(* Logix 5000 project; controller Seperator 1756-L85E rev 33.11; software revision 33.01; part 7 of 7 *)
(* tags used below, declared in another part *)
   Aborted : SFC_STEP;
   Aborting : SFC_STEP;
   Auto_Manual : BOOL;
   CV1 : REAL;
   CV2 : REAL;
   CV3 : DINT;
   Equilibrating : SFC_STEP;
   FI101 : REAL;
   FI102 : REAL;
   FillerPUD1 : RampUpDn;
   FillerPUD2 : RampUpDn;
   FillerPUD3 : RampUpDn;
   FillerPUD4 : RampUpDn;
   FillerPUD5 : RampUpDn;
   FillerPUD6 : RampUpDn;
   FillerPUD7 : RampUpDn;
   Filling : SFC_STEP;
   Flushing : SFC_STEP;
   Half_Sec_PLs : TIMER;
   Holding : SFC_STEP;
   Idle : SFC_STEP;
   II101 : REAL;
   Led_Code : INT;
   LevelUD1 : RampUpDn;
   LI101 : REAL;
   Main_Sequencer : DINT;
   MyP_Motor : P_Motor;   // My (Single-Speed, Non-Reversing) Motor
   PI102 : REAL;
   Qtr_Sec_PLs : TIMER;
   Random : AOI_SIM_RNG_Simple;
   Restarting : SFC_STEP;
   Sec_PLs : TIMER;
   Seperating : SFC_STEP;
   Seperator_Control : PHASE;
   Speeding : SFC_STEP;
   Starting : SFC_STEP;
   Status_Code : INT;
   Stopped : SFC_STEP;
   Stopping : SFC_STEP;
   T1 : FBD_TIMER;
   TI101 : REAL;
   TI101_Temperature : REAL;
   TI101_Temperature_PID_CV : REAL;
   TI101_Temperature_PID_PV : REAL;
   TI101_Temperature_PID_SP : REAL;
   VI101 : REAL;
(* Main_Sequencer, continued *)

ROUTINE Main_Sequencer   (* ladder *)
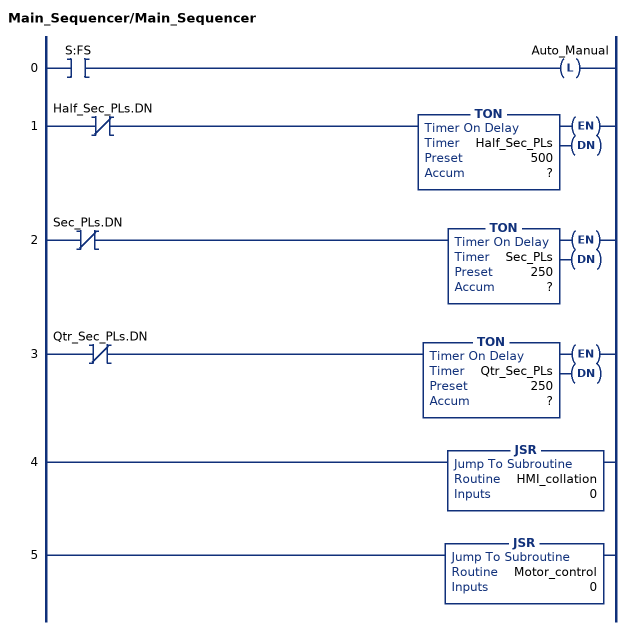
   0: XIC(S:FS)OTL(Auto_Manual);
   1: XIO(Half_Sec_PLs.DN)TON(Half_Sec_PLs,?,?);
   2: XIO(Sec_PLs.DN)TON(Sec_PLs,?,?);
   3: XIO(Qtr_Sec_PLs.DN)TON(Qtr_Sec_PLs,?,?);
   4: JSR(HMI_collation,0);
   5: JSR(Motor_control,0);
END_ROUTINE

ROUTINE Motor_control   (* ladder *)
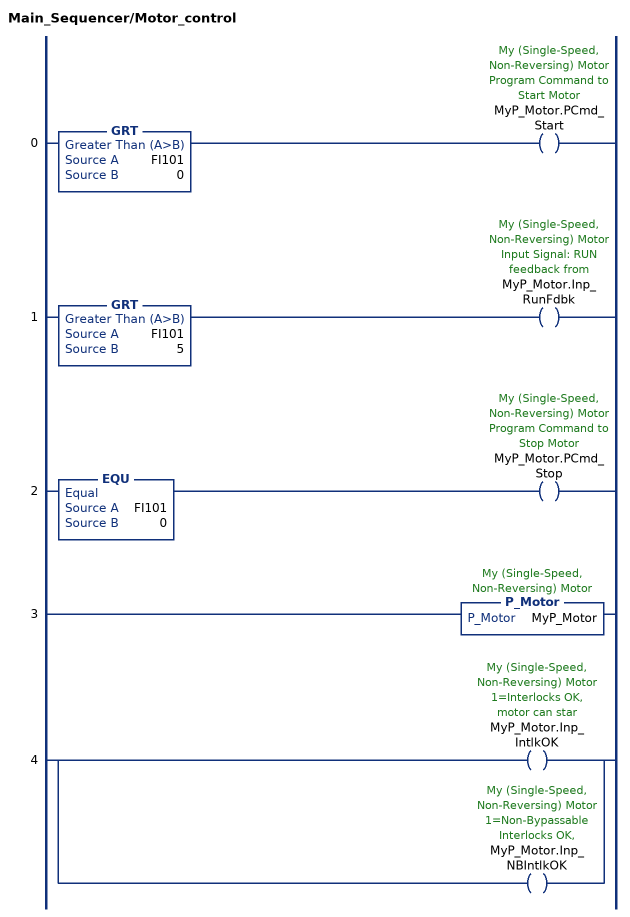
   0: GRT(FI101,0)OTE(MyP_Motor.PCmd_Start);
   1: GRT(FI101,5)OTE(MyP_Motor.Inp_RunFdbk);
   2: EQU(FI101,0)OTE(MyP_Motor.PCmd_Stop);
   3: P_Motor(MyP_Motor);
   4: [OTE(MyP_Motor.Inp_IntlkOK) ,OTE(MyP_Motor.Inp_NBIntlkOK) ];
END_ROUTINE
END_PROGRAM

PROGRAM RandomProgram   (* main routine RandomRoutine *)
VAR
   fsn : REAL := 0.19112337;
END_VAR

ROUTINE RandomRoutine   (* ladder *)
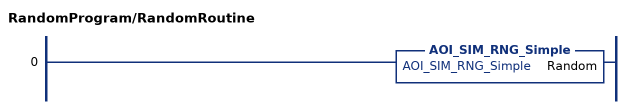
   0: AOI_SIM_RNG_Simple(Random);
END_ROUTINE
END_PROGRAM

PROGRAM RandomUpDown   (* main routine main *)
VAR
   dice001 : AOI_SIM_RNG_Simple := (Seed := 521288629, Count := 470, Number := 0.55877805);
   mult : REAL := 0.025;
   signal : REAL := 0.8641962;
   up : BOOL := 1;
END_VAR

ROUTINE main   (* ladder *)
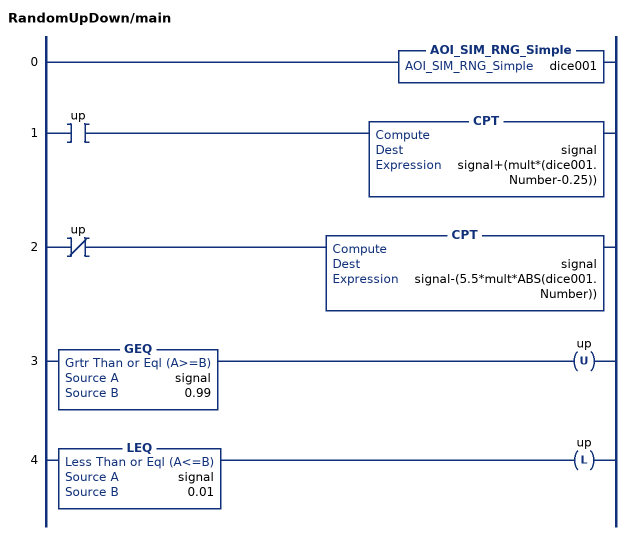
   0: AOI_SIM_RNG_Simple(dice001);
   1: XIC(up)CPT(signal,signal+(mult*(dice001.Number-0.25)));
   2: XIO(up)CPT(signal,signal-(5.5*mult*ABS(dice001.Number)));
   3: GEQ(signal,0.99)OTU(up);
   4: LEQ(signal,0.01)OTL(up);
END_ROUTINE
END_PROGRAM

PROGRAM Seperator_Control
VAR
   Action_000 : SFC_ACTION := (Status := 16#0020_0000, PauseTimer := 1, Count := 1);
   Action_001 : SFC_ACTION := (Status := 16#0020_0000, PauseTimer := 1, Count := 1);
   Action_002 : SFC_ACTION := (Status := 16#0020_0000, PauseTimer := 1, Count := 1);
   Action_003 : SFC_ACTION := (Status := 16#0020_0000, PauseTimer := 1, Count := 1);
   Action_004 : SFC_ACTION := (Status := 16#0020_0000, PauseTimer := 1, Count := 1);
   Action_005 : SFC_ACTION := (Status := 16#0020_0000, PauseTimer := 1, PRE := 5000);
   Action_006 : SFC_ACTION := (Status := 16#0020_0000, PauseTimer := 1, PRE := 5000);
   Action_007 : SFC_ACTION := (Status := 16#0020_0000, PauseTimer := 1, Count := 1);
   Action_008 : SFC_ACTION := (Status := 16#0020_0000, PauseTimer := 1);
   Action_009 : SFC_ACTION := (Status := 16#0020_0000, PauseTimer := 1);
   Action_010 : SFC_ACTION := (Status := 16#0020_0000, PauseTimer := 1, PRE := 5000);
   Action_011 : SFC_ACTION := (Status := 16#0020_0000, PauseTimer := 1);
   Action_012 : SFC_ACTION := (Status := 16#0020_0000, PauseTimer := 1);
   Action_013 : SFC_ACTION := (Status := 16#0020_0000, PauseTimer := 1);
   Action_014 : SFC_ACTION := (Status := 16#0020_0000, PauseTimer := 1);
   Action_015 : SFC_ACTION := (Status := 16#0020_0000, PauseTimer := 1);
   Action_016 : SFC_ACTION := (Status := 16#0020_0000, PauseTimer := 1);
   Action_017 : SFC_ACTION := (Status := 16#0020_0000, PauseTimer := 1, PRE := 5000);
   Action_018 : SFC_ACTION := (Status := 16#0020_0000, PauseTimer := 1);
   Action_019 : SFC_ACTION := (Status := 16#0020_0000, PauseTimer := 1);
   Action_020 : SFC_ACTION := (Status := 16#0020_0000, PauseTimer := 1);
   Action_021 : SFC_ACTION := (Status := 16#0020_0000, PauseTimer := 1);
   Action_022 : SFC_ACTION := (Status := 16#0020_0000, PauseTimer := 1, PRE := 5000);
   Action_023 : SFC_ACTION := (Status := 16#0020_0000, PauseTimer := 1, PRE := 5000);
   Action_024 : SFC_ACTION := (Status := 16#0020_0000, PauseTimer := 1);
   Action_025 : SFC_ACTION := (Status := 16#0020_0000, PauseTimer := 1);
   Action_026 : SFC_ACTION := (Status := 16#0020_0000, PauseTimer := 1, Count := 1);
   Action_027 : SFC_ACTION := (Status := 16#0020_0000, PauseTimer := 1);
   Action_028 : SFC_ACTION := (Status := 16#0020_0000, PauseTimer := 1, Count := 1);
   Breaking : SFC_STEP := (Status := 16#0020_0001, PauseTimer := 1);
   Step_000 : SFC_STEP := (Status := 16#a820_0201, X := 1, SA := 1, DN := 1, PauseTimer := 1, T := 1386790, TMax := 1386790, Count := 2);
   Step_001 : SFC_STEP := (Status := 16#0820_0001, DN := 1, PauseTimer := 1, T := 10, TMax := 10, Count := 1);
   Step_002 : SFC_STEP := (Status := 16#0820_0001, DN := 1, PauseTimer := 1, T := 10, TMax := 10, Count := 1);
   Step_003 : SFC_STEP := (Status := 16#0820_0001, DN := 1, PauseTimer := 1, T := 10, TMax := 10, Count := 1);
   Step_004 : SFC_STEP := (Status := 16#0820_0001, DN := 1, PauseTimer := 1, T := 10, TMax := 10, Count := 1);
   Step_005 : SFC_STEP := (Status := 16#0820_0001, DN := 1, PauseTimer := 1, T := 12950, TMax := 12950, Count := 1);
   Step_006 : SFC_STEP := (Status := 16#0020_0201, PauseTimer := 1);
   Step_007 : SFC_STEP := (Status := 16#0020_0001, PauseTimer := 1);
   Step_008 : SFC_STEP := (Status := 16#0020_0201, PauseTimer := 1);
   Step_009 : SFC_STEP := (Status := 16#0020_0001, PauseTimer := 1);
   Step_010 : SFC_STEP := (Status := 16#a020_0001, X := 1, SA := 1, PauseTimer := 1, PRE := 60000, T := 11750, TMax := 11750, Count := 1);
   Step_011 : SFC_STEP := (Status := 16#0020_0001, PauseTimer := 1);
   Step_012 : SFC_STEP := (Status := 16#0020_0201, PauseTimer := 1);
   Step_013 : SFC_STEP := (Status := 16#0020_0001, PauseTimer := 1);
   Step_014 : SFC_STEP := (Status := 16#0020_0001, PauseTimer := 1);
   Step_015 : SFC_STEP := (Status := 16#0020_0001, PauseTimer := 1);
   Step_016 : SFC_STEP := (Status := 16#0020_0001, PauseTimer := 1);
   Step_017 : SFC_STEP := (Status := 16#0020_0001, PauseTimer := 1);
   Step_018 : SFC_STEP := (Status := 16#0020_0001, PauseTimer := 1);
   Step_019 : SFC_STEP := (Status := 16#0020_0001, PauseTimer := 1);
   Step_020 : SFC_STEP := (Status := 16#0020_0201, PauseTimer := 1);
   Step_021 : SFC_STEP := (Status := 16#0020_0001, PauseTimer := 1);
   Step_022 : SFC_STEP := (Status := 16#0020_0001, PauseTimer := 1);
   Step_023 : SFC_STEP := (Status := 16#0020_0001, PauseTimer := 1);
   Step_024 : SFC_STEP := (Status := 16#0020_0001, PauseTimer := 1, PRE := 120000);
   Stop_000 : SFC_STOP := (Status := 16#0000_2001);
   Stop_001 : SFC_STOP := (Status := 16#0000_2001);
   Stop_002 : SFC_STOP := (Status := 16#0000_2001);
   Stop_003 : SFC_STOP := (Status := 16#0000_2001);
   Stop_004 : SFC_STOP := (Status := 16#0000_2001);
   Tran_000 : BOOL := 1;
   Tran_001 : BOOL := 1;
   Tran_002 : BOOL;
   Tran_003 : BOOL := 1;
   Tran_004 : BOOL := 1;
   Tran_005 : BOOL := 1;
   Tran_006 : BOOL;
   Tran_007 : BOOL;
   Tran_008 : BOOL := 1;
   Tran_009 : BOOL := 1;
   Tran_010 : BOOL;
   Tran_011 : BOOL := 1;
   Tran_012 : BOOL := 1;
   Tran_013 : BOOL := 1;
   Tran_014 : BOOL := 1;
   Tran_015 : BOOL := 1;
   Tran_016 : BOOL := 1;
   Tran_017 : BOOL := 1;
   Tran_018 : BOOL := 1;
   Tran_019 : BOOL := 1;
   Tran_020 : BOOL;
   Tran_021 : BOOL;
   Tran_022 : BOOL;
   Tran_023 : BOOL := 1;
   Tran_024 : BOOL := 1;
   Tran_025 : BOOL := 1;
END_VAR

ROUTINE Aborting   (* sequential function chart *)
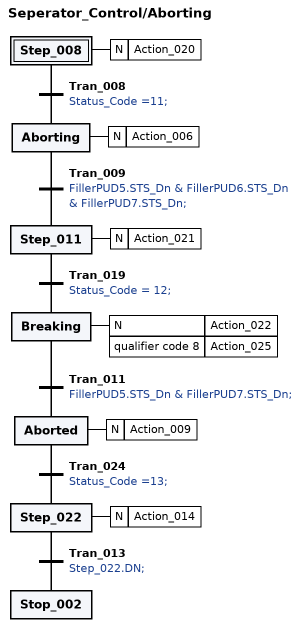
   INITIAL_STEP Step_008:
      ACTION Action_020 (N):
         PI102 :=1.5;
         TI101_Temperature_PID_SP :=56;
         Led_Code := 2;
         Status_Code :=11;
         
         CV1:= FI101;
         CV2:= FI102;
         CV3:= II101;
         
         FillerPUD5.CMD_Start :=0;
         FillerPUD6.CMD_Start :=0;
         FillerPUD7.CMD_Start :=0;
      END_ACTION
   END_STEP
   TRANSITION Tran_008 FROM Step_008 TO Aborting
      := Status_Code =11;
   END_TRANSITION
   STEP Aborting:
      ACTION Action_006 (N):
         //Ramp up the flow and current in 5 seconds
         FillerPUD5.CMD_Start :=1;
         FillerPUD6.CMD_Start :=1;
         FillerPUD7.CMD_Start :=1;
         
         RampUpDn(FillerPUD5,CV1,1,5,FI101);
         RampUpDn(FillerPUD6,CV2,0,5,FI102);
         RampUpDn(FillerPUD7,CV3,7,5,II101);
      END_ACTION
   END_STEP
   TRANSITION Tran_009 FROM Aborting TO Step_011
      := FillerPUD5.STS_Dn & FillerPUD6.STS_Dn & FillerPUD7.STS_Dn;
         
   END_TRANSITION
   STEP Step_011:
      ACTION Action_021 (N):
         Status_Code :=12;
         
         CV1:= VI101;
         CV3:= II101;
         
         FillerPUD5.CMD_Start :=0;
         FillerPUD7.CMD_Start :=0;
      END_ACTION
   END_STEP
   TRANSITION Tran_019 FROM Step_011 TO Breaking
      := Status_Code = 12;
   END_TRANSITION
   STEP Breaking:
      ACTION Action_022 (N):
         //Ramp up the flow and current in 5 seconds
         
         FillerPUD5.CMD_Start :=1;
         FillerPUD7.CMD_Start :=1;
         // if PF755:I.DriveStatus_Active then PF755:O.LogicCommand_Stop :=1; end_if; //Stop seperator
         // PF755:O.Reference :=0;
         
         RampUpDn(FillerPUD1,CV1,0,5,VI101);
         RampUpDn(FillerPUD7,CV3,0,5,II101);
         
         // if PF525:I.Active & PF525_Drive_FP.Sts_ProgramModeEnabled then PF525:O.Stop :=1; end_if; //Stop outlet pump
         
      END_ACTION
      ACTION Action_025 (qualifier code 8):
         // PF755:O.LogicCommand_Stop :=0;
      END_ACTION
   END_STEP
   TRANSITION Tran_011 FROM Breaking TO Aborted
      := FillerPUD5.STS_Dn & FillerPUD7.STS_Dn;
         
   END_TRANSITION
   STEP Aborted:
      ACTION Action_009 (N):
         TI101_Temperature_PID_SP := 20.0;
         PI102 :=0.0;
         FI102 :=0.0;
         Status_Code :=13;
         Led_Code := 1;
      END_ACTION
   END_STEP
   TRANSITION Tran_024 FROM Aborted TO Step_022
      := Status_Code =13;
   END_TRANSITION
   STEP Step_022:
      ACTION Action_014 (N):
         PSC();
      END_ACTION
   END_STEP
   TRANSITION Tran_013 FROM Step_022 TO Stop_002
      := Step_022.DN;
   END_TRANSITION
   STOP Stop_002;
END_ROUTINE

ROUTINE Holding   (* sequential function chart *)
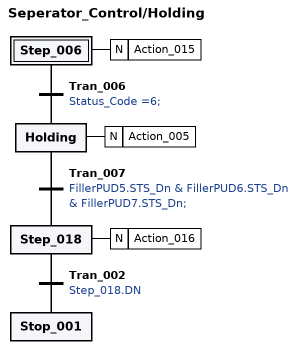
   INITIAL_STEP Step_006:
      ACTION Action_015 (N):
         Led_Code := 2;
         Status_Code :=6;
         PI102 :=1.5;
         CV1:= FI101;
         CV2:= FI102;
         CV3:= II101;
         FillerPUD5.CMD_Start :=0;
         FillerPUD6.CMD_Start :=0;
         FillerPUD7.CMD_Start :=0;
         
      END_ACTION
   END_STEP
   TRANSITION Tran_006 FROM Step_006 TO Holding
      := Status_Code =6;
   END_TRANSITION
   STEP Holding:
      ACTION Action_005 (N):
         //Ramp up the flow and current in 5 seconds
         FillerPUD5.CMD_Start :=1;
         FillerPUD6.CMD_Start :=1;
         FillerPUD7.CMD_Start :=1;
         
         RampUpDn(FillerPUD5,CV1,1,5,FI101);
         RampUpDn(FillerPUD6,CV2,0,5,FI102);
         RampUpDn(FillerPUD7,CV3,7.0,5,II101);
         
      END_ACTION
   END_STEP
   TRANSITION Tran_007 FROM Holding TO Step_018
      := FillerPUD5.STS_Dn & FillerPUD6.STS_Dn & FillerPUD7.STS_Dn;
         
   END_TRANSITION
   STEP Step_018:
      ACTION Action_016 (N):
         Status_Code :=15 ;
         PSC();
         
      END_ACTION
   END_STEP
   TRANSITION Tran_002 FROM Step_018 TO Stop_001
      := Step_018.DN
   END_TRANSITION
   STOP Stop_001;
END_ROUTINE

ROUTINE Resetting   (* structured text *)
   // Reset all the SFC's before returning the phase state to idle
   
   sfr(Aborting,0);
   sfr(Running,0);
   sfr(Holding,0);
   sfr(Stopping,0);
   
   Status_Code :=14;
   Led_Code := 1;
   
   FillerPUD1.CMD_Start :=0;
   FillerPUD2.CMD_Start :=0;
   FillerPUD3.CMD_Start :=0;
   FillerPUD4.CMD_Start :=0;
   FillerPUD5.CMD_Start :=0;
   FillerPUD6.CMD_Start :=0;
   FillerPUD7.CMD_Start :=0;
   
   // if PF755:I.DriveStatus_Active then PF755:O.Reference :=0; end_if;
   // if PF525:I.Active then PF525:O.Stop :=1; end_if;
   
   RampUpDn(FillerPUD1,0.0,0,1,VI101);
   RampUpDn(FillerPUD2,0.0,0,1,II101);
   RampUpDn(FillerPUD3,0.0,0,1,VI101);
   RampUpDn(FillerPUD5,0.0,0,1,FI101);
   RampUpDn(FillerPUD6,0.0,0,1,FI102);
   RampUpDn(FillerPUD7,0.0,0,1,II101);
   
   FI101 :=0.0;
   FI102 :=0.0;
   TI101_Temperature_PID_SP := 20.0;
   PI102 :=0.0;
   II101 :=0.0;
   VI101 := 0;
   
   
   //Wait 30s then change the status to IDLE
   
   T1.PRE :=15000;T1.TimerEnable :=1;
   Tonr(T1);
   if T1.DN then Status_Code :=0; PSC(); end_if;
   
   
   
END_ROUTINE

ROUTINE Restarting   (* sequential function chart *)
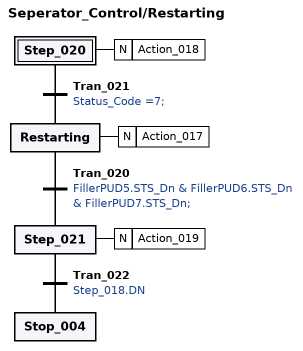
   INITIAL_STEP Step_020:
      ACTION Action_018 (N):
         Led_Code := 3;
         Status_Code :=7;
         
         CV1:= FI101;
         CV2:= FI102;
         CV3:= II101;
         
         FillerPUD5.CMD_Start :=0;
         FillerPUD6.CMD_Start :=0;
         FillerPUD7.CMD_Start :=0;
         
      END_ACTION
   END_STEP
   TRANSITION Tran_021 FROM Step_020 TO Restarting
      := Status_Code =7;
   END_TRANSITION
   STEP Restarting:
      ACTION Action_017 (N):
         //Ramp up the flow and current in 5 seconds
         
         FillerPUD5.CMD_Start :=1;
         FillerPUD6.CMD_Start :=1;
         FillerPUD7.CMD_Start :=1;
         
         RampUpDn(FillerPUD5,CV1,10,5,FI101);
         RampUpDn(FillerPUD6,CV2,8,5,FI102);
         RampUpDn(FillerPUD7,CV3,12,5,II101);
      END_ACTION
   END_STEP
   TRANSITION Tran_020 FROM Restarting TO Step_021
      := FillerPUD5.STS_Dn & FillerPUD6.STS_Dn & FillerPUD7.STS_Dn;
         
   END_TRANSITION
   STEP Step_021:
      ACTION Action_019 (N):
         PSC();
      END_ACTION
   END_STEP
   TRANSITION Tran_022 FROM Step_021 TO Stop_004
      := Step_018.DN
   END_TRANSITION
   STOP Stop_004;
END_ROUTINE

ROUTINE Running   (* sequential function chart *)
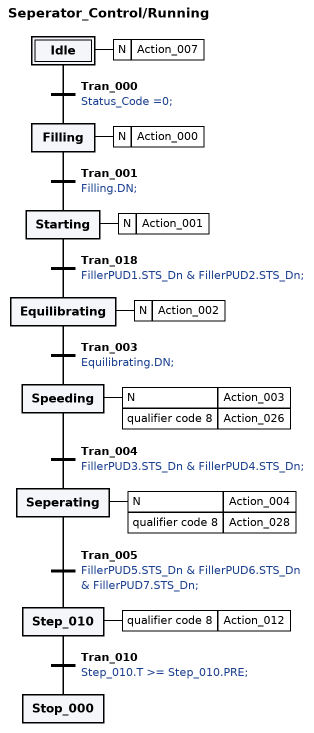
   INITIAL_STEP Idle:
      ACTION Action_007 (N):
         FI101 :=0.0;
         FI102 :=0.0;
         TI101_Temperature_PID_SP := 20.0;
         PI102 :=0.0;
         II101 :=0.0;
         VI101 := 0;
         Led_Code := 1;
         Status_Code :=0;
      END_ACTION
   END_STEP
   TRANSITION Tran_000 FROM Idle TO Filling
      := Status_Code =0;
   END_TRANSITION
   STEP Filling:
      ACTION Action_000 (N):
         FI101 :=1.0;
         TI101_Temperature_PID_SP := 56.0;
         PI102 :=1.0;
         Status_Code :=1;
         Led_Code := 1;
      END_ACTION
   END_STEP
   TRANSITION Tran_001 FROM Filling TO Starting
      := Filling.DN;
   END_TRANSITION
   STEP Starting:
      ACTION Action_001 (N):
         PI102 :=1.5;
         Led_Code := 2;
         Status_Code :=2;
         //Ramp up the speed and current in 5 seconds
         FillerPUD1.CMD_Start :=1;
         FillerPUD2.CMD_Start :=1;
         FillerPUD5.CMD_Start :=1;
         LevelUD1.CMD_Start :=1;
         
         // if not PF755:I.DriveStatus_Active then PF755:O.LogicCommand_Start :=1; end_if; //Start seperator
         // PF755:O.Reference :=10;
         
         RampUpDn(FillerPUD1,0.0,1000,5,VI101);
         RampUpDn(FillerPUD2,0.0,5.0,5,II101);
         RampUpDn(FillerPUD5,1,10,5,FI101);
         
      END_ACTION
   END_STEP
   TRANSITION Tran_018 FROM Starting TO Equilibrating
      := FillerPUD1.STS_Dn & FillerPUD2.STS_Dn;
   END_TRANSITION
   STEP Equilibrating:
      ACTION Action_002 (N):
         Status_Code :=3;
         
         
      END_ACTION
   END_STEP
   TRANSITION Tran_003 FROM Equilibrating TO Speeding
      := Equilibrating.DN;
   END_TRANSITION
   STEP Speeding:
      ACTION Action_003 (N):
         PI102 :=2.0;
         Status_Code :=4;
         
         //Ramp up the speed and current in 5 seconds
         FillerPUD3.CMD_Start :=1;
         FillerPUD4.CMD_Start :=1;
         // if not PF755:I.DriveStatus_Active then PF755:O.LogicCommand_Start :=1;  end_if; //Start seperator
         // PF755:O.Reference :=50;
         RampUpDn(FillerPUD3,1000,5000,5,VI101);
         RampUpDn(FillerPUD4,5,8,5,II101);
         RampUpDn(LevelUD1,20,95,10,LI101);
         
      END_ACTION
      ACTION Action_026 (qualifier code 8):
         // PF755:O.LogicCommand_Start :=0;
      END_ACTION
   END_STEP
   TRANSITION Tran_004 FROM Speeding TO Seperating
      := FillerPUD3.STS_Dn & FillerPUD4.STS_Dn;
         
         
   END_TRANSITION
   STEP Seperating:
      ACTION Action_004 (N):
         Status_Code :=5;
         Led_Code := 3;
         
         
         // if not PF525:I.Active & PF525_Drive_FP.Sts_ProgramModeEnabled then PF525:O.Start :=1; end_if; //Start outlet pump if it is stopped
         
         //Ramp up the flow and current in 5 seconds
         FillerPUD6.CMD_Start :=1;
         FillerPUD7.CMD_Start :=1;
         //Ramp down the tank level
         LevelUD1.CMD_Start :=1;
         
         RampUpDn(FillerPUD6,0,8,5,FI102);
         RampUpDn(FillerPUD7,8,12,5,II101);
         RampUpDn(LevelUD1,95,20,30,LI101);
      END_ACTION
      ACTION Action_028 (qualifier code 8):
         // PF525:O.Start :=0;
      END_ACTION
   END_STEP
   TRANSITION Tran_005 FROM Seperating TO Step_010
      := FillerPUD5.STS_Dn & FillerPUD6.STS_Dn & FillerPUD7.STS_Dn;
         
   END_TRANSITION
   STEP Step_010:
      ACTION Action_012 (qualifier code 8):
         PSC();
      END_ACTION
   END_STEP
   TRANSITION Tran_010 FROM Step_010 TO Stop_000
      := Step_010.T >= Step_010.PRE;
   END_TRANSITION
   STOP Stop_000;
END_ROUTINE

ROUTINE Stopping   (* sequential function chart *)
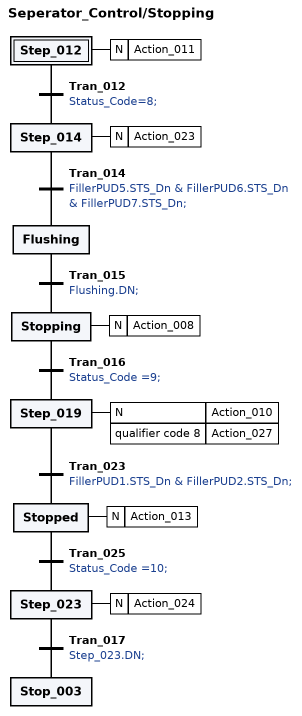
   INITIAL_STEP Step_012:
      ACTION Action_011 (N):
         PI102 :=2;
         TI101 :=56;
         Led_Code := 2;
         Status_Code :=8;
         
         CV1:= FI101;
         CV2:= FI102;
         CV3:= II101;
         
         FillerPUD5.CMD_Start :=0;
         FillerPUD6.CMD_Start :=0;
         FillerPUD7.CMD_Start :=0;
      END_ACTION
   END_STEP
   TRANSITION Tran_012 FROM Step_012 TO Step_014
      := Status_Code=8;
   END_TRANSITION
   STEP Step_014:
      ACTION Action_023 (N):
         //Ramp up the flow and current in 5 seconds
         FillerPUD5.CMD_Start :=1;
         FillerPUD6.CMD_Start :=1;
         FillerPUD7.CMD_Start :=1;
         
         RampUpDn(FillerPUD5,CV1,1,5,FI101);
         RampUpDn(FillerPUD6,CV2,0,5,FI102);
         RampUpDn(FillerPUD7,CV3,7,5,II101);
         
         
      END_ACTION
   END_STEP
   TRANSITION Tran_014 FROM Step_014 TO Flushing
      := FillerPUD5.STS_Dn & FillerPUD6.STS_Dn & FillerPUD7.STS_Dn;
         
   END_TRANSITION
   STEP Flushing:
   END_STEP
   TRANSITION Tran_015 FROM Flushing TO Stopping
      := Flushing.DN;
   END_TRANSITION
   STEP Stopping:
      ACTION Action_008 (N):
         Status_Code :=9;
         
         CV1:= VI101;
         CV2:= II101;
         
         FillerPUD1.CMD_Start :=0;
         FillerPUD2.CMD_Start :=0;
      END_ACTION
   END_STEP
   TRANSITION Tran_016 FROM Stopping TO Step_019
      := Status_Code =9;
         
   END_TRANSITION
   STEP Step_019:
      ACTION Action_010 (N):
         //Ramp up the flow and current in 15 seconds
         FillerPUD1.CMD_Start :=1;
         FillerPUD2.CMD_Start :=1;
         
         // if PF755:I.DriveStatus_Active then PF755:O.LogicCommand_Stop :=1; end_if; //Stop seperator
         
         RampUpDn(FillerPUD1,CV1,0,15,VI101);
         RampUpDn(FillerPUD2,CV2,0,15,II101);
         
         // if PF525:I.Active then PF525:O.Stop :=1; end_if; //Stop outlet pump
      END_ACTION
      ACTION Action_027 (qualifier code 8):
         // PF755:O.LogicCommand_Stop :=0;
         // PF525:O.Stop :=0;
      END_ACTION
   END_STEP
   TRANSITION Tran_023 FROM Step_019 TO Stopped
      := FillerPUD1.STS_Dn & FillerPUD2.STS_Dn;
   END_TRANSITION
   STEP Stopped:
      ACTION Action_013 (N):
         FI101 :=0.0;
         PI102 :=0.0;
         II101 :=0.0;
         Status_Code :=10;
         Led_Code := 4;
         
      END_ACTION
   END_STEP
   TRANSITION Tran_025 FROM Stopped TO Step_023
      := Status_Code =10;
   END_TRANSITION
   STEP Step_023:
      ACTION Action_024 (N):
         PSC();
      END_ACTION
   END_STEP
   TRANSITION Tran_017 FROM Step_023 TO Stop_003
      := Step_023.DN;
   END_TRANSITION
   STOP Stop_003;
END_ROUTINE
END_PROGRAM

PROGRAM TI101_Temperature   (* main routine Initialization *)
VAR
   Amplitude : REAL := 50.0;
   Autotune : PIDE_AUTOTUNE;
   DeadTimeSim : DEADTIME := (Gain := 1.0, RTSTime := 1000, DeltaT := 2.0);
   DEDT_01 : DEADTIME := (Deadtime := 5.0, Gain := 1.4, RTSTime := 1, DeltaT := 0.01, Status := 16#0000_0005, InstructFault := 1, DeadtimeInv := 1);
   DEDT_02 : DEADTIME := (In := 43.287064, Deadtime := 5.0, Gain := 1.4, RTSTime := 1, Out := 60.601887, DeltaT := 0.01, Status := 16#0000_0005, InstructFault := 1, DeadtimeInv := 1);
   DEDT_ARRAY : REAL[1];
   LDLG : LEAD_LAG := (Lag := 55.0, Gain := 1.0, RTSTime := 1, Out := 59.672882, DeltaT := 2.0);
   Temperature_T101 : PID_ENHANCED := (PV := 61.882988, PVEUMax := 300.0, SPProg := 56.0, SPOper := 56.0, SPHLimit := 300.0, RatioProg := 1.0, RatioOper := 1.0, RatioHLimit := 1.0, RatioLLimit := 1.0, CVEUMax := 300.0, CVHLimit := 100.0, PGain := 1.5432097, IGain := 1111.111, DGain := 8.5733875e-05, ProgProgReq := 1, ProgAutoReq := 1, RTSTime := 1000, CVLAlarm := 1, SP := 56.0, SPPercent := 18.666666, PVPercent := 20.627663, E := -5.882988, EPercent := -1.9609966, InitPrimary := 1, WindupLOut := 1, Ratio := 1.0, ProgOper := 1, Auto := 1, DeltaT := 2.0);
   TI101HeateFillerodeAuto : BOOL := 1;
END_VAR

ROUTINE Initialization   (* ladder *)
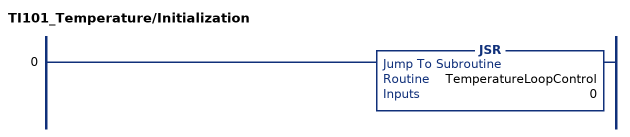
   0: JSR(TemperatureLoopControl,0);
END_ROUTINE

ROUTINE TemperatureLoopControl   (* function block diagram *)
   SHEET 1
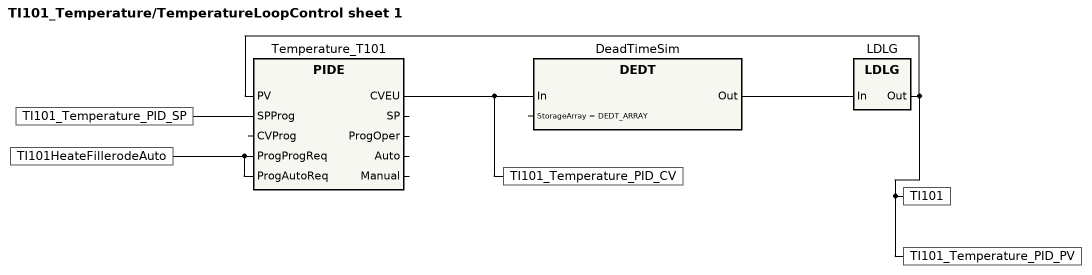
   Temperature_T101 : PIDE(PV := LDLG.Out {feedback}, SPProg := TI101_Temperature_PID_SP, ProgProgReq := TI101HeateFillerodeAuto, ProgAutoReq := TI101HeateFillerodeAuto);   // unwired pins: CVProg SP ProgOper Auto Manual
   TI101_Temperature_PID_CV := Temperature_T101.CVEU;
   DeadTimeSim : DEDT(In := Temperature_T101.CVEU, StorageArray := DEDT_ARRAY);
   LDLG : LDLG(In := DeadTimeSim.Out);
   TI101 := LDLG.Out;
   TI101_Temperature_PID_PV := LDLG.Out;
END_ROUTINE
END_PROGRAM
